
   //-----------------------------------------
   // Enableclosedloop
   //-----------------------------------------
         AN    "DB613_Komponent_State".MeteringPump[4].Enableclosedloop;
         JC    SDA4;
         L     2#0000_0010;
         L     #ControlFlowIndex;
         OW;
         T     #ControlFlowIndex;

   //-----------------------------------------
   // Trigger SDA
   //-----------------------------------------
   SDA4: ON    "DB613_Komponent_State".MeteringPump[4].Puls_SDA;
         O(;
         L     "DB613_Komponent_State".FlowPumpQPB[4];
         L     0.0;
         ==R;
         );
         O(;
         L     "DB613_Komponent_State".PressurePumpQPB[4];
         L     0.0;
         ==R;
         );
         JC    TAB4;
         L     2#0000_1000;
         L     #ControlFlowIndex;
         OW;
         T     #ControlFlowIndex;

   //-----------------------------------------
   // Write Output
   //-----------------------------------------
   TAB4: L     0;
         L     "PN_FlowRate".Component[4].FlowC_F.Address;
         <>D;
         JCN   ed04;
         L     16;
         +D;
         SLD   3;
         LAR1;
         L     #ControlFlowIndex;
         T     PQB [ AR1 , P#0.0 ];

   //----------------------------------------------------------------
   // Tandem comand
   //----------------------------------------------------------------
   ta04: NOP   0;
   //      L     0
   //      L     "DB1233_ProCanIO_Flow".AddressFlow[4].Ref_TandemComand
   //      <I
   //      SPBN  ed01
   //      SLD   3
   //      LAR1
   //
   //      CALL  BLKMOV
   //         blk_type:=Any
   //         SRCBLK  :="DB206_TandemCommand".PistonPair[4]
   //         RET_VAL :=#TemRetBLKMOV
   //         DSTBLK  :=#TempTandem
   //
   //      L     #TempTandem
   //      TAW
   //      T PAB [ AR1 , P#0.0 ]

   ed04: NOP   0;
END_REGION

REGION Network 5: Common conditions production mode mixinghead
   // Service/Production mixinghead machine 1
         A     "DB619_State_MPart".Operationmode[1].Operation;
         AN    "DB619_State_MPart".ShotMa[1].ShotData.ShotDisabled;
         A     "DB619_State_MPart".Operationmode[1].Auto;
         AN    "DB619_State_MPart".Operationmode[1].Test;
         =     #TempShotWithMaterial_M1;

   // Service/Production mixinghead machine 2
         A     "DB619_State_MPart".Operationmode[2].Operation;
         AN    "DB619_State_MPart".ShotMa[2].ShotData.ShotDisabled;
         A     "DB619_State_MPart".Operationmode[2].Auto;
         AN    "DB619_State_MPart".Operationmode[2].Test;
         =     #TempShotWithMaterial_M2;
END_REGION

REGION Network 6
         L     "GetToolShotValues_DB".IO_PartShotNoNew;
         T     "ShotNoNextMa1";

         AN    "DB619_State_MPart".Cycle[1].running;
         R     "StopShotCorrMH01";
         R     "StopShotCorrMH02";
         R     "StopShotCorrMH03";
         R     "StopShotCorrMH04";
         R     "StopShotCorrMH05";
         R     "StopShotCorrMH06";
         R     "StopShotCorrMH07";
         R     "StopShotCorrMH08";
END_REGION

REGION Network 7: Mixinghead 1
   //--- mixinghead 1 active at a machine ----------------
         O(;
         L     "DB619_State_MPart".ShotMa[1].ShotData.MH_No;
         L     1;
         ==I;
         );
         O(;
         L     "DB619_State_MPart".ShotMa[2].ShotData.MH_No;
         L     1;
         ==I;
         );
         =     #Temp_MH_Shot_MH01;
         JCN   cr01;

         L     "DB704_MH_Value".Mixinghead[1].Corrvalue;
         T     #Temp_CorrValue;

   // Shottime correction
   cr01: NOP   0;
   //----------------------------------------------------------------
   // Read Shottime for next shot
   //----------------------------------------------------------------
         O     "DB619_State_MPart".Cycle[1].PressurizeTimeRuns;
         O     "DB619_State_MPart".Cycle[1].CtrlChangeTimeRuns;
         A     #Temp_MH_Shot_MH01;
         =     "F_CycleRunningMH01";  // Read corr Shottime

         A     #Temp_MH_Shot_MH01;
         A     "DB619_State_MPart".SWU[1].SWU_OK;
         JCN   om01;

         A     "DB619_State_MPart".Operationmode[1].Operation;
         AN    "DB619_State_MPart".ShotMa[1].ShotData.ShotDisabled;
         =     #Temp_OperationMode;

         AN    "DB619_State_MPart".Cycle[1].running;
         R     "StopShotCorrMH01";
         A     "DB110_Interf_Program_M1".Bits.Stop_Cycle;
         A     "DB619_State_MPart".Cycle[1].running;
         S     "StopShotCorrMH01";

         O     "StopShotCorrMH01";
         O     "DB009_Faults".Fault_State_Grp_1_M1;
         ON    "DB619_State_MPart".Operationmode[1].Controllvoltage;
         =     #Temp_Error;

         CALL  "FC215_SHOT_ADJUST"
         ( IN_Cycle_running   := "F_CycleRunningMH01",
           IN_Shot_running    := "M_ShotActive",
           IN_OP_Mode_foaming := #Temp_OperationMode,
           IN_Error_GRP_1     := #Temp_Error,
           IN_Tool_no         := "DB619_State_MPart".ToolMa[1].ToolNo,
           IN_PS_no           := "ShotNoNextMa1",
           IN_Set_Shottime_DB := "DB606_PV_Machine".Machine[1].ShotTime.PV_SetV.Value,
           IN_Actual_Shottime := "DB606_PV_Machine".Machine[1].ShotTime.PV_ActV.Value,
           IN_Corrvalue       := #Temp_CorrValue,
           IN_DB_Shotadjust   := "DB315_ShotadjustS",
           IN_ShotRelease     := "DB619_State_MPart".Cycle[1].Shotrelease,
           IN_MhManual        := 0,  //"DB123_MH_IO_Signals".MH[1].IN.MH_Manual_Mode
           IO_Correct_factor  := "DB614_MH_State".ShotAdjustMH[1].CorrFact,
           IO_PAD_Shottime    := "DB614_MH_State".ShotAdjustMH[1].FoamingTime_ProCan,
           IO_Modul_activ     := "DB614_MH_State".ShotAdjustMH[1].ShotCorrActive,
           IO_Helpflag        := "DB614_MH_State".ShotAdjustMH[1].HFShotCorr,
           IO_Last_Shottime   := "DB614_MH_State".ShotAdjustMH[1].LastShottime,
           IO_Soll_for_Corr   := "DB614_MH_State".ShotAdjustMH[1].SetValueForCorr,
           IO_AdrCorrF        := "DB614_MH_State".ShotAdjustMH[1].AdrCorrFact,
           IO_TestProgram     := "DB614_MH_State".ShotAdjustMH[1].ShotCorrTest,
           IO_CorrTimeTest    := "DB614_MH_State".ShotAdjustMH[1].CorrTimeTest
         );

   // Write mixinghead data to procan mudule
   //----------------------------------------------------------------------
   // Check if the communication partner is ready for
   // data transfer to ProCan
   // ---------------------------------------------------------------------
   om01: NOP   0;
         AN    "PN_Mixinghead".Mixinghead[1].Digital.Active;
         AN    "PN_Mixinghead".Mixinghead[1].Analog.Active;
         JC    em01;

   //-----------------------------------------------------------------
   // Output signals of mixing head modul 1
   //-----------------------------------------------------------------

   //    L     "DB1232_ProCanIO_MH".AddressMH[1].Ref_Digital_Input
   //    L     16
   //    >D
   //    SPB   MD01
   //    U     "DB123_MH_IO_Signals".MH[1].OUT.MH.H_CP_Back_MH
   //    =     "H_CP_Back_MH1"
   //    U     "DB123_MH_IO_Signals".MH[1].OUT.MH.H_Rel_Foaming_MH
   //    =     "H_Rel_Foaming_MH1"
   //    U     "DB123_MH_IO_Signals".MH[1].OUT.MH.H_HighPressure_MH
   //    =     "H_HighPressure_MH1"
   //    U     "DB123_MH_IO_Signals".MH[1].OUT.MH.K_Fault_MC
   //    =     "K_Stoerung_FT"
   //    U     "DB123_MH_IO_Signals".MH[1].OUT.MH.K_ShotEnd_MC
   //    =     "K_Schussende_FT"
   //    U     "DB123_MH_IO_Signals".MH[1].OUT.MH.V_MH
   //    =     "V_MH_open_MH1"
   //    U     "DB123_MH_IO_Signals".MH[1].OUT.MH.V_CP_Forward_MH
   //    =     "V_CP_Forward_MH1"
   //    SPA   MH01


   MD01: NOP   0;

         A     "DB123_MH_IO_Signals".MH[1].OUT.MH.V_SWU_MH;
         =     "V_SWU_MH01";
         A     "DB123_MH_IO_Signals".MH[1].OUT.MH.H_Shotcounter_MH;
         =     "H_Shotcounter_MH01";

         A     "DB704_MH_Value".Mixinghead[1].Cleaning_Piston.ContrCleaningPiston;
         JC    nocp;
         A     "DB123_MH_IO_Signals".MH[1].OUT.MH.V_CP_Forward_MH;
         =     "V_CP_Forward_MH01";

   nocp: A     "DB123_MH_IO_Signals".MH[1].OUT.MH.H_CP_Back_MH;
         =     "H_CP_Back_MH01";

         A     "DB123_MH_IO_Signals".MH[1].OUT.MH.H_Rel_Foaming_MH;
         =     "H_Rel_Foaming_MH01";
         A     "DB123_MH_IO_Signals".MH[1].OUT.MH.H_HighPressure_MH;
         =     "H_HighPressure_MH01";
         A     "DB123_MH_IO_Signals".MH[1].OUT.MH.K_Fault_MC;
         =     "K_Fault_MC01";
         A     "DB123_MH_IO_Signals".MH[1].OUT.MH.K_ShotEnd_MC;
         =     "K_ShotEnd_MC01";
         A     "DB123_MH_IO_Signals".MH[1].OUT.MH.V_MH;
         =     "V_MH_open_MH01";
         A     "DB123_MH_IO_Signals".MH[1].OUT.MH.V_LowPressure_Circ_MH;
         =     "V_LowPressure_Circ_MH01";

   //------------------------------------------------------------
   //
   //     Activate mixinghead at ProCan  modul
   //
   //------------------------------------------------------------

   //--------------- Mixinghead 1--------------------------------
   MH01: O     #Temp_MH_Shot_MH01;
         JCN   SV01;

   //-----------------------------------------------------------------
   // Transmit calculated shot time to ProCan
   //-----------------------------------------------------------------
         L     0;
         L     "PN_Mixinghead".Mixinghead[1].Digital.Address;
         <>D;
         JCN   SV01;
         SLD   3;
         LAR1;
         L     "DB614_MH_State".ShotAdjustMH[1].FoamingTime_ProCan;
         T     PQD [ AR1 , P#0.0 ];
   SV01: NOP   0;

   //*****************************************************************
   // Shot control of mixing head
   //*****************************************************************
         L     0;
         T     #ControlBitShot;
   //--------------------------------------------------
   // Shotcycle finished reset signals
   //--------------------------------------------------
         AN    "DB619_State_MPart".Mixinghead[1].Mixingheadvalve."01";
         R     "ShotFinishedModul_MH01";
         R     "EnableFinishShot_MH01";

   //-------------------------------------------------
   //  Signal enable shot finish  101.12.HK
   //-------------------------------------------------
         O(;
   //    u    LastBreakFromExternal    // Signal vom ROBOTER !!!
         A     "DB123_MH_IO_Signals".MH[1].IN.MH_Status.shotactive_MH;
         );
         ON    "DB704_MH_Value".Mixinghead[1].ShotBreak;
         O     "DB123_MH_IO_Signals".MH[1].IN.MH_Manual_Mode;
         S     "EnableFinishShot_MH01";

   //-------------------------------------------------
   // Signal to reset shotrelease
   //-------------------------------------------------
         ON    "DB123_MH_IO_Signals".MH[1].IN.MH_Status.shotactive_MH;
         O     "EnableFinishShot_MH01";
         A     "DB123_MH_IO_Signals".MH[1].IN.MH_Status.shotdone_MH;
         S     "ShotFinishedModul_MH01";

   //-------------------------------------------------
   // Shot release
   //-------------------------------------------------
         A     "DB619_State_MPart".Mixinghead[1].Mixingheadvalve."01";
         AN    "ShotFinishedModul_MH01";
         AN    "DB009_Faults".Fault_State_Grp_1_M1;
         AN    "DB009_Faults".Faults_FKT_Grp_1_M1;
         JCN   SO01;
         L     2#0000_0001;
         L     #ControlBitShot;
         OW;
         T     #ControlBitShot;
   //-------------------------------------------------
   // Shot without Timer
   //-------------------------------------------------
   SO01: CLR;
         JCN   SW01;
         L     2#0000_0010;
         L     #ControlBitShot;
         OW;
         T     #ControlBitShot;
   //-------------------------------------------------
   // Shot with Timer
   //-------------------------------------------------
   SW01: A     "DB619_State_MPart".Mixinghead[1].Mixingheadvalve."01";
         AN    "ShotFinishedModul_MH01";
         AN    "DB009_Faults".Fault_State_Grp_1_M1;
         AN    "DB009_Faults".Faults_FKT_Grp_1_M1;
         JCN   SP01;
         L     2#0000_0100;
         L     #ControlBitShot;
         OW;
         T     #ControlBitShot;
   //-----------------------------------------------------------------
   // Service / Production
   //-----------------------------------------------------------------
   SP01: NOP   0;
         A(;
         ON    #TempShotWithMaterial_M1;
         ON    "DB619_State_MPart".MH_at_Machine[1]."01";
         );
         A(;
         ON    #TempShotWithMaterial_M2;
         ON    "DB619_State_MPart".MH_at_Machine[2]."01";
         );
         AN    "DB619_State_MPart".Operationmode[1].Test;
         ON    "DB614_MH_State".MH_Status[1].Switch_Service_ON_OFF;
         JCN   RF01;
         L     2#0000_1000;
         L     #ControlBitShot;
         OW;
         T     #ControlBitShot;
   //-----------------------------------------------------------------
   // Spare Bit 4..6
   //-----------------------------------------------------------------

   //-----------------------------------------------------------------
   // Reset faults
   //-----------------------------------------------------------------
   RF01: A     "DB009_Faults".HF_Faults_Quit;  // "DB009_Faults".Faults_Reset_FKT_M1
         JCN   FE01;
         L     2#1000_0000;
         L     #ControlBitShot;
         OW;
         T     #ControlBitShot;

   FE01: NOP   0;
   //-----------------------------------------------------------------
   // Write Output MH Status
   //-----------------------------------------------------------------
         L     "PN_Mixinghead".Mixinghead[1].Digital.Address;
         L     4;
         +D;
         SLD   3;
         LAR1;
         L     #ControlBitShot;
         T     PQB [ AR1 , P#0.0 ];
   //*****************************************************************
   // Cleaning Piston control of mixing head
   //*****************************************************************
         L     0;
         T     #ControlBitCP;
   //-----------------------------------
   // Request cleaning piston after shot
   //-----------------------------------
         A     "DB619_State_MPart".ShotMa[1].ShotData.CP_AfterShot;
   //    U     "DB704_MH_Value".Mixinghead[1].WithCleaningPiston
         JCN   CF01;
         L     2#0000_0001;
         L     #ControlBitCP;
         OW;
         T     #ControlBitCP;
   //-----------------------------------
   // Request cleaning piston with button
   //-----------------------------------
   CF01: A     "DB614_MH_State".MH_CleaningPiston[1].CP_valve_selected;
         JCN   CM01;
         L     2#0000_0010;
         L     #ControlBitCP;
         OW;
         T     #ControlBitCP;
   //-----------------------------------
   // Break forward time
   //-----------------------------------
   CM01: NOP   0;

   //-----------------------------------------------------------------
   // Reset faults
   //-----------------------------------------------------------------
         A     "DB009_Faults".HF_Faults_Quit;
         JCN   FC01;
         L     2#0000_1000;
         L     #ControlBitCP;
         OW;
         T     #ControlBitCP;

   FC01: NOP   0;
   //-----------------------------------------------------------------
   // Write Output CP Status
   //-----------------------------------------------------------------
         L     0;
         L     "PN_Mixinghead".Mixinghead[1].ReinigungskolbenDigital.Address;
         <>D;
         JCN   em01;
         SLD   3;
         LAR1;
         L     #ControlBitCP;
         T     PQB [ AR1 , P#0.0 ];

         JU    em01;

   //*****************************************************************
   // Setvalue position of cleaning piston MH 1
   //*****************************************************************
   //      L     "DB896_ConfAnaCP_Contr".AnaCleaningPiston[1].RearPosition
   //      UN    "DB610_State_MPart".Cycle_Ma[1].running
   //      SPB   gap1
   //      L     "DB610_State_MPart".ShotMa[1].ShotValues.CP_ThrottleGap
   //      ITD
   //      DTR
   //      L     "DB604_PV_Mixinghead".Mixinghead[1].CleaningPiston.PV_Conf_ActV.Multiplier
   //      *R
   //      RND
   //      L     "DB604_PV_Mixinghead".Mixinghead[1].CleaningPiston.PV_Conf_ActV.OffsetSignal
   //      ITD
   //      +D
   //gap1: T     #ThrottleGap
   //
   //      L     0
   //      L     "DB1232_ProCanIO_MH".AddressMH[1].Ref_PLC_set_value_CP
   //      <D
   //      SPBN  nz01
   //      SLD   3
   //      LAR1
   //      L     #ThrottleGap
   //      T PAW [ AR1 , P#0.0 ]


   //*******************************************************************
   // Nozzel control of mixing head 1
   //*******************************************************************
   nz01: L     0;  // Bei 0 immer Bypass
   //     T     #TempNozzelBitCirc
   //
   //     L     "DB704_MH_Value".Mixinghead[1].NozzelShot
   //     T     #TempNozzelBitShot
   //
   //     L     0
   //     L     "DB1232_ProCanIO_MH".AddressMH[1].Ref_NozzelBypassControl
   //     <D
   //     SPBN  fr01
   //     SLD   3
   //     LAR1
   //     L     #TempNozzelBitShot
   //     T PAB [ AR1 , P#0.0 ]
   //
   //      L     #TempNozzelBitCirc
   //      T PAB [ AR1 , P#1.0 ]
   //
   //-----------------------------------------------------------------
   // Nozzel/bypass force  mixing head 1
   //-----------------------------------------------------------------
   //fr01: L     "DB704_MH_Value".Mixinghead[1].NozzelForcen
   //      T     #TempNozzelBitForce
   //
   //      L     "DB704_MH_Value".Mixinghead[1].NozzleRelease
   //      T     #TempNozzelBitRelease
   //
   //      L     0
   //      L     "DB1232_ProCanIO_MH".AddressMH[1].Ref_NozzelBypassSetOut
   //      <D
   //      SPBN  em01
   //      SLD   3
   //      LAR1
   //      L     #TempNozzelBitForce
   //      T PAB [ AR1 , P#0.0 ]
   //
   //      L     #TempNozzelBitRelease
   //      T PAB [ AR1 , P#1.0 ]
   //
   em01: NOP   0;
END_REGION

REGION Network 8: Mixinghead 2
   //--- mixinghead 2 active at a machine ----------------
         O(;
         L     "DB619_State_MPart".ShotMa[1].ShotData.MH_No;
         L     2;
         ==I;
         );
         O(;
         L     "DB619_State_MPart".ShotMa[2].ShotData.MH_No;
         L     2;
         ==I;
         );
         =     #Temp_MH_Shot_MH02;
         JCN   cr02;

         L     "DB704_MH_Value".Mixinghead[2].Corrvalue;
         T     #Temp_CorrValue;

   // Shottime correction
   cr02: NOP   0;

   //----------------------------------------------------------------
   // Read Shottime for next shot
   //----------------------------------------------------------------
         O     "DB619_State_MPart".Cycle[1].PressurizeTimeRuns;
         O     "DB619_State_MPart".Cycle[1].CtrlChangeTimeRuns;
         A     #Temp_MH_Shot_MH02;
         =     "F_CycleRunningMH02";  // Read corr Shottime

         A     #Temp_MH_Shot_MH02;
         A     "DB619_State_MPart".SWU[1].SWU_OK;
         JCN   om02;

         A     "DB619_State_MPart".Operationmode[1].Operation;
         AN    "DB619_State_MPart".ShotMa[1].ShotData.ShotDisabled;
         =     #Temp_OperationMode;

         A     "DB110_Interf_Program_M1".Bits.Stop_Cycle;
         A     "DB619_State_MPart".Cycle[1].running;
         S     "StopShotCorrMH02";

         O     "StopShotCorrMH02";
         O     "DB009_Faults".Fault_State_Grp_1_M1;
         ON    "DB619_State_MPart".Operationmode[1].Controllvoltage;
   //      ON    "DB123_MH_IO_Signals".MH[2].IN.MH_Status.shotdone_MH
         =     #Temp_Error;


         CALL  "FC215_SHOT_ADJUST"
         ( IN_Cycle_running   := "F_CycleRunningMH02",  // "DB610_State_MPart".Cycle_Ma[1].running
           IN_Shot_running    := "M_ShotActive",
           IN_OP_Mode_foaming := #Temp_OperationMode,
           IN_Error_GRP_1     := #Temp_Error,
           IN_Tool_no         := "DB619_State_MPart".ToolMa[1].ToolNo,
           IN_PS_no           := "ShotNoNextMa1",
           IN_Set_Shottime_DB := "DB606_PV_Machine".Machine[1].ShotTime.PV_SetV.Value,
           IN_Actual_Shottime := "DB606_PV_Machine".Machine[1].ShotTime.PV_ActV.Value,
           IN_Corrvalue       := #Temp_CorrValue,
           IN_DB_Shotadjust   := "DB315_ShotadjustS",
           IN_ShotRelease     := "DB619_State_MPart".Cycle[1].Shotrelease,
           IN_MhManual        := 0,  //"DB123_MH_IO_Signals".MH[2].IN.MH_Manual_Mode
           IO_Correct_factor  := "DB614_MH_State".ShotAdjustMH[2].CorrFact,
           IO_PAD_Shottime    := "DB614_MH_State".ShotAdjustMH[2].FoamingTime_ProCan,
           IO_Modul_activ     := "DB614_MH_State".ShotAdjustMH[2].ShotCorrActive,
           IO_Helpflag        := "DB614_MH_State".ShotAdjustMH[2].HFShotCorr,
           IO_Last_Shottime   := "DB614_MH_State".ShotAdjustMH[2].LastShottime,
           IO_Soll_for_Corr   := "DB614_MH_State".ShotAdjustMH[2].SetValueForCorr,
           IO_AdrCorrF        := "DB614_MH_State".ShotAdjustMH[2].AdrCorrFact,
           IO_TestProgram     := "DB614_MH_State".ShotAdjustMH[2].ShotCorrTest,
           IO_CorrTimeTest    := "DB614_MH_State".ShotAdjustMH[2].CorrTimeTest
         );

   // Write mixinghead data to procan mudule
   //----------------------------------------------------------------------
   // Check if the communication partner is ready for
   // data transfer to ProCan
   // ---------------------------------------------------------------------
   om02: NOP   0;
         AN    "PN_Mixinghead".Mixinghead[2].Digital.Active;
         AN    "PN_Mixinghead".Mixinghead[2].Analog.Active;
         JC    em02;
   //-----------------------------------------------------------------
   // Output signals of mixing head modul 2
   //-----------------------------------------------------------------
         A     "DB123_MH_IO_Signals".MH[2].OUT.MH.V_SWU_MH;
         =     "V_SWU_MH02";
         A     "DB123_MH_IO_Signals".MH[2].OUT.MH.H_Shotcounter_MH;
         =     "H_Shotcounter_MH02";
         A     "DB123_MH_IO_Signals".MH[2].OUT.MH.V_CP_Forward_MH;
         =     "V_CP_Forward_MH02";
         A     "DB123_MH_IO_Signals".MH[2].OUT.MH.H_CP_Back_MH;
         =     "H_CP_Back_MH02";
         A     "DB123_MH_IO_Signals".MH[2].OUT.MH.H_Rel_Foaming_MH;
         =     "H_Rel_Foaming_MH02";
         A     "DB123_MH_IO_Signals".MH[2].OUT.MH.H_HighPressure_MH;
         =     "H_HighPressure_MH02";
         A     "DB123_MH_IO_Signals".MH[2].OUT.MH.K_Fault_MC;
         =     "K_Fault_MC02";
         A     "DB123_MH_IO_Signals".MH[2].OUT.MH.K_ShotEnd_MC;
         =     "K_ShotEnd_MC02";
         A     "DB123_MH_IO_Signals".MH[2].OUT.MH.V_MH;
         =     "V_MH_open_MH02";
         A     "DB123_MH_IO_Signals".MH[2].OUT.MH.V_LowPressure_Circ_MH;
         =     "V_LowPressure_Circ_MH02";

   //------------------------------------------------------------
   //
   //     Activate mixinghead at ProCan  modul
   //
   //------------------------------------------------------------

   //--------------- Mixinghead 2--------------------------------
         O     #Temp_MH_Shot_MH02;
         JCN   SV02;
   //-----------------------------------------------------------------
   // Transmit calculated shot time to ProCan
   //-----------------------------------------------------------------
         L     0;
         L     "PN_Mixinghead".Mixinghead[2].Digital.Address;
         <>D;
         JCN   SV02;
         SLD   3;
         LAR1;
         L     "DB614_MH_State".ShotAdjustMH[2].FoamingTime_ProCan;
         T     PQD[AR1, P#0.0];
   SV02: NOP   0;

   //*****************************************************************
   // Shot control of mixing head
   //*****************************************************************
         L     0;
         T     #ControlBitShot;
   //--------------------------------------------------
   // Shotcycle finished reset signals
   //--------------------------------------------------
         AN    "DB619_State_MPart".Mixinghead[1].Mixingheadvalve."02";
         R     "ShotFinishedModul_MH02";
         R     "EnableFinishShot_MH02";

   //-------------------------------------------------
   //  Signal enable shot finish
   //-------------------------------------------------
         O(;
   //    u    LastBreakFromExternal    // Signal vom ROBOTER !!!
         A     "DB123_MH_IO_Signals".MH[2].IN.MH_Status.shotactive_MH;
         );
         ON    "DB704_MH_Value".Mixinghead[2].ShotBreak;
         O     "DB123_MH_IO_Signals".MH[2].IN.MH_Manual_Mode;
         S     "EnableFinishShot_MH02";

   //-------------------------------------------------
   // Signal to reset shotrelease
   //-------------------------------------------------
         ON    "DB123_MH_IO_Signals".MH[2].IN.MH_Status.shotactive_MH;
         O     "EnableFinishShot_MH02";
         A     "DB123_MH_IO_Signals".MH[2].IN.MH_Status.shotdone_MH;
         S     "ShotFinishedModul_MH02";
   //-------------------------------------------------
   // Shot release
   //-------------------------------------------------
         A     "DB619_State_MPart".Mixinghead[1].Mixingheadvalve."02";
         AN    "ShotFinishedModul_MH02";
         AN    "DB009_Faults".Fault_State_Grp_1_M1;
         AN    "DB009_Faults".Faults_FKT_Grp_1_M1;
         JCN   SO02;
         L     2#0000_0001;
         L     #ControlBitShot;
         OW;
         T     #ControlBitShot;
   //-------------------------------------------------
   // Shot without Timer
   //-------------------------------------------------
   SO02: CLR;
         JCN   SW02;
         L     2#0000_0010;
         L     #ControlBitShot;
         OW;
         T     #ControlBitShot;
   //-------------------------------------------------
   // Shot with Timer
   //-------------------------------------------------
   SW02: A     "DB619_State_MPart".Mixinghead[1].Mixingheadvalve."02";
         AN    "ShotFinishedModul_MH02";
         AN    "DB009_Faults".Fault_State_Grp_1_M1;
         AN    "DB009_Faults".Faults_FKT_Grp_1_M1;
         JCN   SP02;
         L     2#0000_0100;
         L     #ControlBitShot;
         OW;
         T     #ControlBitShot;
   //-----------------------------------------------------------------
   // Service / Production
   //-----------------------------------------------------------------
   SP02: NOP   0;
         A(;
         ON    #TempShotWithMaterial_M1;
         ON    "DB619_State_MPart".MH_at_Machine[1]."02";
         );
         A(;
         ON    #TempShotWithMaterial_M2;
         ON    "DB619_State_MPart".MH_at_Machine[2]."02";
         );
         ON    "DB614_MH_State".MH_Status[2].Switch_Service_ON_OFF;
         JCN   RF02;
         L     2#0000_1000;
         L     #ControlBitShot;
         OW;
         T     #ControlBitShot;

   //-----------------------------------------------------------------
   // Spare Bit 4..6
   //-----------------------------------------------------------------

   //-----------------------------------------------------------------
   // Reset faults
   //-----------------------------------------------------------------
   RF02: A     "DB009_Faults".HF_Faults_Quit;
         JCN   FE02;
         L     2#1000_0000;
         L     #ControlBitShot;
         OW;
         T     #ControlBitShot;

   FE02: NOP   0;
   //-----------------------------------------------------------------
   // Write Output MH Status
   //-----------------------------------------------------------------
         L     "PN_Mixinghead".Mixinghead[2].Digital.Address;
         L     4;
         +D;
         SLD   3;
         LAR1;
         L     #ControlBitShot;
         T     PQB [ AR1 , P#0.0 ];
   //*****************************************************************
   // Cleaning Piston control of mixing head
   //*****************************************************************
         O(;
         L     "PN_Mixinghead".Mixinghead[2].ReinigungskolbenDigital.Address;
         L     0;
         ==I;
         );
         ON    "PN_Mixinghead".Mixinghead[2].ReinigungskolbenDigital.Active;
         JC    em02;

         L     0;
         T     #ControlBitCP;
   //-------------------------------------------------
   // Request cleaning piston after shot
   //-------------------------------------------------
         A     "DB619_State_MPart".ShotMa[1].ShotData.CP_AfterShot;
   //    U     "DB704_MH_Value".Mixinghead[1].WithCleaningPiston
         JCN   CF02;
         L     2#0000_0001;
         L     #ControlBitCP;
         OW;
         T     #ControlBitCP;
   //-------------------------------------------------
   // Request cleaning piston with button
   //-------------------------------------------------
   CF02: A     "DB614_MH_State".MH_CleaningPiston[2].CP_valve_selected;
         JCN   CM02;
         L     2#0000_0010;
         L     #ControlBitCP;
         OW;
         T     #ControlBitCP;
   //-------------------------------------------------
   // Break forward time
   //-------------------------------------------------
   CM02: NOP   0;
   //-----------------------------------------------------------------
   // Reset faults
   //-----------------------------------------------------------------
         A     "DB009_Faults".HF_Faults_Quit;
         JCN   FC02;
         L     2#0000_1000;
         L     #ControlBitCP;
         OW;
         T     #ControlBitCP;
   //-------------------------------------------------
   FC02: NOP   0;
   //-------------------------------------------------
   // Write Output CP Status
   //-------------------------------------------------
         L     "PN_Mixinghead".Mixinghead[2].ReinigungskolbenDigital.Address;
         SLD   3;
         LAR1;
         L     #ControlBitCP;
         T     PQB [ AR1 , P#0.0 ];
   //-------------------------------------------------
         JU    em02;
   //*****************************************************************
   // Setvalue position of cleaning piston MH 2
   //*****************************************************************
   //      L     "DB896_ConfAnaCP_Contr".AnaCleaningPiston[2].RearPosition
   //      UN    "DB610_State_MPart".Cycle_Ma[1].running
   //      SPB   gap1
   //      L     "DB610_State_MPart".ShotMa[1].ShotValues.CP_ThrottleGap
   //      ITD
   //      DTR
   //      L     "DB604_PV_Mixinghead".Mixinghead[2].CleaningPiston.PV_Conf_ActV.Multiplier
   //      *R
   //      RND
   //      L     "DB604_PV_Mixinghead".Mixinghead[2].CleaningPiston.PV_Conf_ActV.OffsetSignal
   //      ITD
   //      +D
   //gap1: T     #ThrottleGap
   //
   //      L     0
   //      L     "DB1232_ProCanIO_MH".AddressMH[2].Ref_PLC_set_value_CP
   //      <D
   //      SPBN  nz01
   //      SLD   3
   //      LAR1
   //      L     #ThrottleGap
   //      T PAW [ AR1 , P#0.0 ]
   em02: NOP   0;
END_REGION

REGION Network 9: Mixinghead 3
   //--- mixinghead 3 active at a machine ----------------
         O(;
         L     "DB619_State_MPart".ShotMa[1].ShotData.MH_No;
         L     3;
         ==I;
         );
         O(;
         L     "DB619_State_MPart".ShotMa[2].ShotData.MH_No;
         L     3;
         ==I;
         );
         =     #Temp_MH_Shot_MH03;
         JCN   cr03;

         L     "DB704_MH_Value".Mixinghead[3].Corrvalue;
         T     #Temp_CorrValue;

   // Shottime correction
   cr03: NOP   0;

   //----------------------------------------------------------------
   // Read Shottime for next shot
   //----------------------------------------------------------------
         O     "DB619_State_MPart".Cycle[1].PressurizeTimeRuns;
         O     "DB619_State_MPart".Cycle[1].CtrlChangeTimeRuns;
         A     #Temp_MH_Shot_MH03;
         =     "F_CycleRunningMH03";  // Read corr Shottime

         A     #Temp_MH_Shot_MH03;
         A     "DB619_State_MPart".SWU[1].SWU_OK;
         JCN   om03;

         A     "DB619_State_MPart".Operationmode[1].Operation;
         AN    "DB619_State_MPart".ShotMa[1].ShotData.ShotDisabled;
         =     #Temp_OperationMode;

         AN    "DB619_State_MPart".Cycle[1].running;
         R     "StopShotCorrMH03";
         A     "DB110_Interf_Program_M1".Bits.Stop_Cycle;
         A     "DB619_State_MPart".Cycle[1].running;
         S     "StopShotCorrMH03";

         O     "StopShotCorrMH03";
         O     "DB009_Faults".Fault_State_Grp_1_M1;
         ON    "DB619_State_MPart".Operationmode[1].Controllvoltage;
   //      ON    "DB123_MH_IO_Signals".MH[3].IN.MH_Status.shotdone_MH

         =     #Temp_Error;

         CALL  "FC215_SHOT_ADJUST"
         ( IN_Cycle_running   := "F_CycleRunningMH03",  // "DB610_State_MPart".Cycle_Ma[1].running
           IN_Shot_running    := "M_ShotActive",
           IN_OP_Mode_foaming := #Temp_OperationMode,
           IN_Error_GRP_1     := #Temp_Error,
           IN_Tool_no         := "DB619_State_MPart".ToolMa[1].ToolNo,
           IN_PS_no           := "ShotNoNextMa1",
           IN_Set_Shottime_DB := "DB606_PV_Machine".Machine[1].ShotTime.PV_SetV.Value,
           IN_Actual_Shottime := "DB606_PV_Machine".Machine[1].ShotTime.PV_ActV.Value,
           IN_Corrvalue       := #Temp_CorrValue,
           IN_DB_Shotadjust   := "DB315_ShotadjustS",
           IN_ShotRelease     := "DB619_State_MPart".Cycle[1].Shotrelease,
           IN_MhManual        := 0,  //"DB123_MH_IO_Signals".MH[3].IN.MH_Manual_Mode
           IO_Correct_factor  := "DB614_MH_State".ShotAdjustMH[3].CorrFact,
           IO_PAD_Shottime    := "DB614_MH_State".ShotAdjustMH[3].FoamingTime_ProCan,
           IO_Modul_activ     := "DB614_MH_State".ShotAdjustMH[3].ShotCorrActive,
           IO_Helpflag        := "DB614_MH_State".ShotAdjustMH[3].HFShotCorr,
           IO_Last_Shottime   := "DB614_MH_State".ShotAdjustMH[3].LastShottime,
           IO_Soll_for_Corr   := "DB614_MH_State".ShotAdjustMH[3].SetValueForCorr,
           IO_AdrCorrF        := "DB614_MH_State".ShotAdjustMH[3].AdrCorrFact,
           IO_TestProgram     := "DB614_MH_State".ShotAdjustMH[3].ShotCorrTest,
           IO_CorrTimeTest    := "DB614_MH_State".ShotAdjustMH[3].CorrTimeTest
         );

   // Write mixinghead data to procan mudule
   //----------------------------------------------------------------------
   // Check if the communication partner is ready for
   // data transfer to ProCan
   // ---------------------------------------------------------------------
   om03: NOP   0;
         AN    "PN_Mixinghead".Mixinghead[3].Digital.Active;
         AN    "PN_Mixinghead".Mixinghead[3].Analog.Active;
         JC    em03;
   //-----------------------------------------------------------------
   // Output signals of mixing head modul 3
   //-----------------------------------------------------------------
         A     "DB123_MH_IO_Signals".MH[3].OUT.MH.V_SWU_MH;
         =     "V_SWU_MH03";
         A     "DB123_MH_IO_Signals".MH[3].OUT.MH.H_Shotcounter_MH;
         =     "H_Shotcounter_MH03";
         A     "DB123_MH_IO_Signals".MH[3].OUT.MH.V_CP_Forward_MH;
         =     "V_CP_Forward_MH03";
         A     "DB123_MH_IO_Signals".MH[3].OUT.MH.H_CP_Back_MH;
         =     "H_CP_Back_MH03";
         A     "DB123_MH_IO_Signals".MH[3].OUT.MH.H_Rel_Foaming_MH;
         =     "H_Rel_Foaming_MH03";
         A     "DB123_MH_IO_Signals".MH[3].OUT.MH.H_HighPressure_MH;
         =     "H_HighPressure_MH03";
         A     "DB123_MH_IO_Signals".MH[3].OUT.MH.K_Fault_MC;
         =     "K_Fault_MC03";
         A     "DB123_MH_IO_Signals".MH[3].OUT.MH.K_ShotEnd_MC;
         =     "K_ShotEnd_MC03";
         A     "DB123_MH_IO_Signals".MH[3].OUT.MH.V_MH;
         =     "V_MH_open_MH03";
   //      U     "DB123_MH_IO_Signals".MH[3].OUT.MH.V_LowPressure_Circ_MH
   //      =     "V_LowPressure_Circ_MH03"

   //------------------------------------------------------------
   //
   //     Activate mixinghead at ProCan  modul
   //
   //------------------------------------------------------------

   //--------------- Mixinghead 3--------------------------------
         O     #Temp_MH_Shot_MH03;
         JCN   SV03;
   //-----------------------------------------------------------------
   // Transmit calculated shot time to ProCan
   //-----------------------------------------------------------------
         L     0;
         L     "PN_Mixinghead".Mixinghead[3].Digital.Address;
         <>D;
         JCN   SV03;
         SLD   3;
         LAR1;
         L     "DB614_MH_State".ShotAdjustMH[3].FoamingTime_ProCan;
         T     PQD[AR1, P#0.0];
   SV03: NOP   0;

   //*****************************************************************
   // Shot control of mixing head
   //*****************************************************************
         L     0;
         T     #ControlBitShot;
   //--------------------------------------------------
   // Shotcycle finished reset signals
   //--------------------------------------------------
         AN    "DB619_State_MPart".Mixinghead[1].Mixingheadvalve."03";
         R     "ShotFinishedModul_MH03";
         R     "EnableFinishShot_MH03";

   //-------------------------------------------------
   //  Signal enable shot finish
   //-------------------------------------------------
         O(;
   //    u    LastBreakFromExternal    // Signal vom ROBOTER !!!
         A     "DB123_MH_IO_Signals".MH[3].IN.MH_Status.shotactive_MH;
         );
         ON    "DB704_MH_Value".Mixinghead[3].ShotBreak;
         O     "DB123_MH_IO_Signals".MH[3].IN.MH_Manual_Mode;
         S     "EnableFinishShot_MH03";

   //-------------------------------------------------
   // Signal to reset shotrelease
   //-------------------------------------------------
         ON    "DB123_MH_IO_Signals".MH[3].IN.MH_Status.shotactive_MH;
         O     "EnableFinishShot_MH03";
         A     "DB123_MH_IO_Signals".MH[3].IN.MH_Status.shotdone_MH;
         S     "ShotFinishedModul_MH03";
   //-------------------------------------------------
   // Shot release
   //-------------------------------------------------
         A     "DB619_State_MPart".Mixinghead[1].Mixingheadvalve."03";
         AN    "ShotFinishedModul_MH03";
         AN    "DB009_Faults".Fault_State_Grp_1_M1;
         AN    "DB009_Faults".Faults_FKT_Grp_1_M1;
         JCN   SO03;
         L     2#0000_0001;
         L     #ControlBitShot;
         OW;
         T     #ControlBitShot;
   //-------------------------------------------------
   // Shot without Timer
   //-------------------------------------------------
   SO03: CLR;
         JCN   SW03;
         L     2#0000_0010;
         L     #ControlBitShot;
         OW;
         T     #ControlBitShot;
   //-------------------------------------------------
   // Shot with Timer
   //-------------------------------------------------
   SW03: A     "DB619_State_MPart".Mixinghead[1].Mixingheadvalve."03";
         AN    "ShotFinishedModul_MH03";
         AN    "DB009_Faults".Fault_State_Grp_1_M1;
         AN    "DB009_Faults".Faults_FKT_Grp_1_M1;
         JCN   SP03;
         L     2#0000_0100;
         L     #ControlBitShot;
         OW;
         T     #ControlBitShot;
   //-----------------------------------------------------------------
   // Service / Production
   //-----------------------------------------------------------------
   SP03: NOP   0;
         A(;
         ON    #TempShotWithMaterial_M1;
         ON    "DB619_State_MPart".MH_at_Machine[1]."03";
         );
         A(;
         ON    #TempShotWithMaterial_M2;
         ON    "DB619_State_MPart".MH_at_Machine[2]."03";
         );
         ON    "DB614_MH_State".MH_Status[3].Switch_Service_ON_OFF;
         JCN   RF03;
         L     2#0000_1000;
         L     #ControlBitShot;
         OW;
         T     #ControlBitShot;
   //-----------------------------------------------------------------
   // Spare Bit 4..6
   //-----------------------------------------------------------------

   //-----------------------------------------------------------------
   // Reset faults
   //-----------------------------------------------------------------
   RF03: A     "DB009_Faults".HF_Faults_Quit;
         JCN   FE03;
         L     2#1000_0000;
         L     #ControlBitShot;
         OW;
         T     #ControlBitShot;

   FE03: NOP   0;
   //-----------------------------------------------------------------
   // Write Output MH Status
   //-----------------------------------------------------------------
         L     "PN_Mixinghead".Mixinghead[3].Digital.Address;
         L     4;
         +D;
         SLD   3;
         LAR1;
         L     #ControlBitShot;
         T     PQB [ AR1 , P#0.0 ];
   //*****************************************************************
   // Cleaning Piston control of mixing head
   //*****************************************************************
         O(;
         L     "PN_Mixinghead".Mixinghead[3].ReinigungskolbenDigital.Address;
         L     0;
         ==I;
         );
         ON    "PN_Mixinghead".Mixinghead[3].ReinigungskolbenDigital.Active;
         JC    em03;

         L     0;
         T     #ControlBitCP;
   //-------------------------------------------------
   // Request cleaning piston after shot
   //-------------------------------------------------
         A     "DB619_State_MPart".ShotMa[1].ShotData.CP_AfterShot;
   //    U     "DB704_MH_Value".Mixinghead[3].WithCleaningPiston
         JCN   CF03;
         L     2#0000_0001;
         L     #ControlBitCP;
         OW;
         T     #ControlBitCP;
   //-------------------------------------------------
   // Request cleaning piston with button
   //-------------------------------------------------
   CF03: A     "DB614_MH_State".MH_CleaningPiston[3].CP_valve_selected;
         JCN   CM03;
         L     2#0000_0010;
         L     #ControlBitCP;
         OW;
         T     #ControlBitCP;
   //-------------------------------------------------
   // Break forward time
   //-------------------------------------------------
   CM03: NOP   0;
   //-----------------------------------------------------------------
   // Reset faults
   //-----------------------------------------------------------------
         A     "DB009_Faults".HF_Faults_Quit;
         JCN   FC03;
         L     2#0000_1000;
         L     #ControlBitCP;
         OW;
         T     #ControlBitCP;
   //-------------------------------------------------
   FC03: NOP   0;
   //-------------------------------------------------
   // Write Output CP Status
   //-------------------------------------------------
         L     "PN_Mixinghead".Mixinghead[3].ReinigungskolbenDigital.Address;
         SLD   3;
         LAR1;
         L     #ControlBitCP;
         T     PQB [ AR1 , P#0.0 ];
   //-------------------------------------------------
         JU    em03;
   //*****************************************************************
   // Setvalue position of cleaning piston MH 3
   //*****************************************************************
   //      L     "DB896_ConfAnaCP_Contr".AnaCleaningPiston[3].RearPosition
   //      UN    "DB610_State_MPart".Cycle_Ma[1].running
   //      SPB   gap1
   //      L     "DB610_State_MPart".ShotMa[1].ShotValues.CP_ThrottleGap
   //      ITD
   //      DTR
   //      L     "DB604_PV_Mixinghead".Mixinghead[3].CleaningPiston.PV_Conf_ActV.Multiplier
   //      *R
   //      RND
   //      L     "DB604_PV_Mixinghead".Mixinghead[3].CleaningPiston.PV_Conf_ActV.OffsetSignal
   //      ITD
   //      +D
   //gap1: T     #ThrottleGap
   //
   //      L     0
   //      L     "DB1232_ProCanIO_MH".AddressMH[3].Ref_PLC_set_value_CP
   //      <D
   //      SPBN  nz01
   //      SLD   3
   //      LAR1
   //      L     #ThrottleGap
   //      T PAW [ AR1 , P#0.0 ]
   //*****************************************************************
   em03: NOP   0;
END_REGION

REGION Network 10: Mixinghead 4
   //--- mixinghead 4 active at a machine ----------------
         O(;
         L     "DB619_State_MPart".ShotMa[1].ShotData.MH_No;
         L     4;
         ==I;
         );
         O(;
         L     "DB619_State_MPart".ShotMa[2].ShotData.MH_No;
         L     4;
         ==I;
         );
         =     #Temp_MH_Shot_MH04;
         JCN   cr04;

         L     "DB704_MH_Value".Mixinghead[4].Corrvalue;
         T     #Temp_CorrValue;

   // Shottime correction
   cr04: NOP   0;

   //----------------------------------------------------------------
   // Read Shottime for next shot
   //----------------------------------------------------------------
         O     "DB619_State_MPart".Cycle[1].PressurizeTimeRuns;
         O     "DB619_State_MPart".Cycle[1].CtrlChangeTimeRuns;
         A     #Temp_MH_Shot_MH04;
         =     "F_CycleRunningMH04";  // Read corr Shottime

         A     #Temp_MH_Shot_MH04;
         A     "DB619_State_MPart".SWU[1].SWU_OK;
         JCN   om04;

         A     "DB619_State_MPart".Operationmode[1].Operation;
         AN    "DB619_State_MPart".ShotMa[1].ShotData.ShotDisabled;
         =     #Temp_OperationMode;

         AN    "DB619_State_MPart".Cycle[1].running;
         R     "StopShotCorrMH04";
         A     "DB110_Interf_Program_M1".Bits.Stop_Cycle;
         A     "DB619_State_MPart".Cycle[1].running;
         S     "StopShotCorrMH04";

         O     "StopShotCorrMH04";
         O     "DB009_Faults".Fault_State_Grp_1_M1;
         ON    "DB619_State_MPart".Operationmode[1].Controllvoltage;
   //      ON    "DB123_MH_IO_Signals".MH[4].IN.MH_Status.shotdone_MH
         =     #Temp_Error;

         CALL  "FC215_SHOT_ADJUST"
         ( IN_Cycle_running   := "F_CycleRunningMH04",  // "DB610_State_MPart".Cycle_Ma[1].running
           IN_Shot_running    := "M_ShotActive",  // "DB610_State_MPart".Cycle_Ma[1].ShotRuns
           IN_OP_Mode_foaming := #Temp_OperationMode,  // "DB610_State_MPart".Operationmode_Ma[1].Operation
           IN_Error_GRP_1     := #Temp_Error,  // "M1001_FaultLevel_1"
           IN_Tool_no         := "DB619_State_MPart".ToolMa[1].ToolNo,
           IN_PS_no           := "ShotNoNextMa1",  // "DB610_State_MPart".ShotDataMa[1].ShotNo
           IN_Set_Shottime_DB := "DB606_PV_Machine".Machine[1].ShotTime.PV_SetV.Value,
           IN_Actual_Shottime := "DB606_PV_Machine".Machine[1].ShotTime.PV_ActV.Value,
           IN_Corrvalue       := #Temp_CorrValue,
           IN_DB_Shotadjust   := "DB315_ShotadjustS",
           IN_ShotRelease     := "DB619_State_MPart".Cycle[1].Shotrelease,
           IN_MhManual        := 0,  //"DB123_MH_IO_Signals".MH[4].IN.MH_Manual_Mode
           IO_Correct_factor  := "DB614_MH_State".ShotAdjustMH[4].CorrFact,
           IO_PAD_Shottime    := "DB614_MH_State".ShotAdjustMH[4].FoamingTime_ProCan,
           IO_Modul_activ     := "DB614_MH_State".ShotAdjustMH[4].ShotCorrActive,
           IO_Helpflag        := "DB614_MH_State".ShotAdjustMH[4].HFShotCorr,
           IO_Last_Shottime   := "DB614_MH_State".ShotAdjustMH[4].LastShottime,
           IO_Soll_for_Corr   := "DB614_MH_State".ShotAdjustMH[4].SetValueForCorr,
           IO_AdrCorrF        := "DB614_MH_State".ShotAdjustMH[4].AdrCorrFact,
           IO_TestProgram     := "DB614_MH_State".ShotAdjustMH[4].ShotCorrTest,
           IO_CorrTimeTest    := "DB614_MH_State".ShotAdjustMH[4].CorrTimeTest
         );

   // Write mixinghead data to procan mudule
   //----------------------------------------------------------------------
   // Check if the communication partner is ready for
   // data transfer to ProCan
   // ---------------------------------------------------------------------
   om04: NOP   0;
         AN    "PN_Mixinghead".Mixinghead[4].Digital.Active;
         AN    "PN_Mixinghead".Mixinghead[4].Analog.Active;
         JC    em04;
   //-----------------------------------------------------------------
   // Output signals of mixing head modul 4
   //-----------------------------------------------------------------
         A     "DB123_MH_IO_Signals".MH[4].OUT.MH.V_SWU_MH;
         =     "V_SWU_MH04";
         A     "DB123_MH_IO_Signals".MH[4].OUT.MH.H_Shotcounter_MH;
         =     "H_Shotcounter_MH04";
         A     "DB123_MH_IO_Signals".MH[4].OUT.MH.V_CP_Forward_MH;
         =     "V_CP_Forward_MH04";
         A     "DB123_MH_IO_Signals".MH[4].OUT.MH.H_CP_Back_MH;
         =     "H_CP_Back_MH04";
         A     "DB123_MH_IO_Signals".MH[4].OUT.MH.H_Rel_Foaming_MH;
         =     "H_Rel_Foaming_MH04";
         A     "DB123_MH_IO_Signals".MH[4].OUT.MH.H_HighPressure_MH;
         =     "H_HighPressure_MH04";
         A     "DB123_MH_IO_Signals".MH[4].OUT.MH.K_Fault_MC;
         =     "K_Fault_MC04";
         A     "DB123_MH_IO_Signals".MH[4].OUT.MH.K_ShotEnd_MC;
         =     "K_ShotEnd_MC04";
         A     "DB123_MH_IO_Signals".MH[4].OUT.MH.V_MH;
         =     "V_MH_open_MH04";
         A     "DB123_MH_IO_Signals".MH[4].OUT.MH.V_LowPressure_Circ_MH;
         =     "V_LowPressure_Circ_MH04";

   //------------------------------------------------------------
   //
   //     Activate mixinghead at ProCan  modul
   //
   //------------------------------------------------------------

   //--------------- Mixinghead 4 --------------------------------
         O     #Temp_MH_Shot_MH04;
         JCN   SV04;

   //-----------------------------------------------------------------
   // Transmit calculated shot time to ProCan
   //-----------------------------------------------------------------
         L     0;
         L     "PN_Mixinghead".Mixinghead[4].Digital.Address;
         <>D;
         JCN   SV04;
         SLD   3;
         LAR1;
         L     "DB614_MH_State".ShotAdjustMH[4].FoamingTime_ProCan;
         T     PQD[AR1, P#0.0];
   SV04: NOP   0;

   //*****************************************************************
   // Shot control of mixing head
   //*****************************************************************
         L     0;
         T     #ControlBitShot;
   //--------------------------------------------------
   // Shotcycle finished reset signals
   //--------------------------------------------------
         AN    "DB619_State_MPart".Mixinghead[1].Mixingheadvalve."04";
         R     "ShotFinishedModul_MH04";
         R     "EnableFinishShot_MH04";

